   5080: 'Carrier 79 Drive: Short-circuit/ground fault detected', class No Acknowledgement, trigger "DB302_HMI_Faults_Carrier79_Faults_1" bit 7
   5081: 'Carrier 79 Drive: PROFINET Setpoint timeout', class No Acknowledgement, trigger "DB302_HMI_Faults_Carrier79_Faults_1" bit 8
   5082: 'Carrier 79 Power unit: Overcurrent', class No Acknowledgement, trigger "DB302_HMI_Faults_Carrier79_Faults_1" bit 9
   5083: 'Carrier 79 Power unit: DC link voltage overvoltage', class No Acknowledgement, trigger "DB302_HMI_Faults_Carrier79_Faults_1" bit 10
   5084: 'Carrier 79 Power unit: DC link voltage undervoltage', class No Acknowledgement, trigger "DB302_HMI_Faults_Carrier79_Faults_1" bit 11
   5085: 'Carrier 79 Power unit: Line phase failure in main circuit', class No Acknowledgement, trigger "DB302_HMI_Faults_Carrier79_Faults_1" bit 12
   5086: 'Carrier 79 Power unit: Phase failure motor cable', class No Acknowledgement, trigger "DB302_HMI_Faults_Carrier79_Faults_1" bit 13
   5087: 'Carrier 79 Power unit: Ground fault', class No Acknowledgement, trigger "DB302_HMI_Faults_Carrier79_Faults_1" bit 14
   5088: 'Spare_Fault_5088', class No Acknowledgement, trigger "DB302_HMI_Faults_Carrier79_Faults_1" bit 15
   5089: 'Carrier 79 Motion Off Fault', class No Acknowledgement, trigger "DB302_HMI_Faults_Carrier79_Faults_2" bit 0
   5090: 'Carrier 79 Motion On Fault', class No Acknowledgement, trigger "DB302_HMI_Faults_Carrier79_Faults_2" bit 1
   5091: 'Carrier 79 Spacing Fault', class No Acknowledgement, trigger "DB302_HMI_Faults_Carrier79_Faults_2" bit 2
   5092: 'Carrier 79 Duplicate Carrier Number Fault', class No Acknowledgement, trigger "DB302_HMI_Faults_Carrier79_Faults_2" bit 3
   5093: 'Spare_Fault_5093', class No Acknowledgement, trigger "DB302_HMI_Faults_Carrier79_Faults_2" bit 4
   5094: 'Spare_Fault_5094', class No Acknowledgement, trigger "DB302_HMI_Faults_Carrier79_Faults_2" bit 5
   5095: 'Spare_Fault_5095', class No Acknowledgement, trigger "DB302_HMI_Faults_Carrier79_Faults_2" bit 6
   5096: 'Spare_Fault_5096', class No Acknowledgement, trigger "DB302_HMI_Faults_Carrier79_Faults_2" bit 7
   5097: 'Spare_Fault_5097', class No Acknowledgement, trigger "DB302_HMI_Faults_Carrier79_Faults_2" bit 8
   5098: 'Spare_Fault_5098', class No Acknowledgement, trigger "DB302_HMI_Faults_Carrier79_Faults_2" bit 9
   5099: 'Spare_Fault_5099', class No Acknowledgement, trigger "DB302_HMI_Faults_Carrier79_Faults_2" bit 10
   5100: 'Spare_Fault_5100', class No Acknowledgement, trigger "DB302_HMI_Faults_Carrier79_Faults_2" bit 11
   5101: 'Spare_Fault_5101', class No Acknowledgement, trigger "DB302_HMI_Faults_Carrier79_Faults_2" bit 12
   5102: 'Spare_Fault_5102', class No Acknowledgement, trigger "DB302_HMI_Faults_Carrier79_Faults_2" bit 13
   5103: 'Spare_Fault_5103', class No Acknowledgement, trigger "DB302_HMI_Faults_Carrier79_Faults_2" bit 14
   5104: 'Spare_Fault_5104', class No Acknowledgement, trigger "DB302_HMI_Faults_Carrier79_Faults_2" bit 15
   5105: 'Spare_Fault_5105', class No Acknowledgement, trigger "DB302_HMI_Faults_Carrier79_Faults_3" bit 0
   5106: 'Spare_Fault_5106', class No Acknowledgement, trigger "DB302_HMI_Faults_Carrier79_Faults_3" bit 1
   5107: 'Spare_Fault_5107', class No Acknowledgement, trigger "DB302_HMI_Faults_Carrier79_Faults_3" bit 2
   5108: 'Spare_Fault_5108', class No Acknowledgement, trigger "DB302_HMI_Faults_Carrier79_Faults_3" bit 3
   5109: 'Spare_Fault_5109', class No Acknowledgement, trigger "DB302_HMI_Faults_Carrier79_Faults_3" bit 4
   5110: 'Spare_Fault_5110', class No Acknowledgement, trigger "DB302_HMI_Faults_Carrier79_Faults_3" bit 5
   5111: 'Spare_Fault_5111', class No Acknowledgement, trigger "DB302_HMI_Faults_Carrier79_Faults_3" bit 6
   5112: 'Spare_Fault_5112', class No Acknowledgement, trigger "DB302_HMI_Faults_Carrier79_Faults_3" bit 7
   5113: 'Spare_Fault_5113', class No Acknowledgement, trigger "DB302_HMI_Faults_Carrier79_Faults_3" bit 8
   5114: 'Spare_Fault_5114', class No Acknowledgement, trigger "DB302_HMI_Faults_Carrier79_Faults_3" bit 9
   5115: 'Spare_Fault_5115', class No Acknowledgement, trigger "DB302_HMI_Faults_Carrier79_Faults_3" bit 10
   5116: 'Spare_Fault_5116', class No Acknowledgement, trigger "DB302_HMI_Faults_Carrier79_Faults_3" bit 11
   5117: 'Spare_Fault_5117', class No Acknowledgement, trigger "DB302_HMI_Faults_Carrier79_Faults_3" bit 12
   5118: 'Spare_Fault_5118', class No Acknowledgement, trigger "DB302_HMI_Faults_Carrier79_Faults_3" bit 13
   5119: 'Spare_Fault_5119', class No Acknowledgement, trigger "DB302_HMI_Faults_Carrier79_Faults_3" bit 14
   5120: 'Spare_Fault_5120', class No Acknowledgement, trigger "DB302_HMI_Faults_Carrier79_Faults_3" bit 15
   5121: 'Carrier 80 Disconnect Open Power Fault DI11.0', class No Acknowledgement, trigger "DB302_HMI_Faults_Carrier80_Faults_0" bit 0
   5122: 'Carrier 80 Drive Profinet Comm Fault', class No Acknowledgement, trigger "DB302_HMI_Faults_Carrier80_Faults_0" bit 1
   5123: 'Carrier 80 Production Stop Not Reset', class No Acknowledgement, trigger "DB302_HMI_Faults_Carrier80_Faults_0" bit 2
   5124: 'Carrier 80 CB02122 Tripped', class No Acknowledgement, trigger "DB302_HMI_Faults_Carrier80_Faults_0" bit 3
   5125: 'Carrier 80 CB02123 Tripped', class No Acknowledgement, trigger "DB302_HMI_Faults_Carrier80_Faults_0" bit 4
   5126: 'Carrier 80 AUX1 CB Tripped', class No Acknowledgement, trigger "DB302_HMI_Faults_Carrier80_Faults_0" bit 5
   5127: 'Carrier 80 AUX2 CB Tripped', class No Acknowledgement, trigger "DB302_HMI_Faults_Carrier80_Faults_0" bit 6
   5128: 'Carrier 80 PLC Not Communicating', class No Acknowledgement, trigger "DB302_HMI_Faults_Carrier80_Faults_0" bit 7
   5129: 'Carrier 80 Safe Input Card Fault', class No Acknowledgement, trigger "DB302_HMI_Faults_Carrier80_Faults_0" bit 8
   5130: 'Carrier 80 Safe Output Card Fault', class No Acknowledgement, trigger "DB302_HMI_Faults_Carrier80_Faults_0" bit 9
   5131: 'Carrier 80 Standard Input Card Fault', class No Acknowledgement, trigger "DB302_HMI_Faults_Carrier80_Faults_0" bit 10
   5132: 'Carrier 80 Standard Output Card Fault', class No Acknowledgement, trigger "DB302_HMI_Faults_Carrier80_Faults_0" bit 11
   5133: 'Carrier 80 Encoder Position Fault', class No Acknowledgement, trigger "DB302_HMI_Faults_Carrier80_Faults_0" bit 12
   5134: 'Carrier 80 Encoder Internal Error', class No Acknowledgement, trigger "DB302_HMI_Faults_Carrier80_Faults_0" bit 13
   5135: 'Carrier 80 Encoder Comm Fault', class No Acknowledgement, trigger "DB302_HMI_Faults_Carrier80_Faults_0" bit 14
   5136: 'Carrier 80 HMI Comm Fault', class No Acknowledgement, trigger "DB302_HMI_Faults_Carrier80_Faults_0" bit 15
   5137: 'Carrier 80 Crash Detection Fault', class No Acknowledgement, trigger "DB302_HMI_Faults_Carrier80_Faults_1" bit 0
   5138: 'Carrier 80 Carrier Number Invalid', class No Acknowledgement, trigger "DB302_HMI_Faults_Carrier80_Faults_1" bit 1
   5139: 'Carrier 80 Drive: PROFINET configuration error', class No Acknowledgement, trigger "DB302_HMI_Faults_Carrier80_Faults_1" bit 2
   5140: 'Carrier 80 Drive: Error internal communications', class No Acknowledgement, trigger "DB302_HMI_Faults_Carrier80_Faults_1" bit 3
   5141: 'Carrier 80 Drive: Motor overtemperature', class No Acknowledgement, trigger "DB302_HMI_Faults_Carrier80_Faults_1" bit 4
   5142: 'Carrier 80 Drive: Motor overcurrent', class No Acknowledgement, trigger "DB302_HMI_Faults_Carrier80_Faults_1" bit 5
   5143: 'Carrier 80 Drive: Infeed or power unit not ready', class No Acknowledgement, trigger "DB302_HMI_Faults_Carrier80_Faults_1" bit 6
   5144: 'Carrier 80 Drive: Short-circuit/ground fault detected', class No Acknowledgement, trigger "DB302_HMI_Faults_Carrier80_Faults_1" bit 7
   5145: 'Carrier 80 Drive: PROFINET Setpoint timeout', class No Acknowledgement, trigger "DB302_HMI_Faults_Carrier80_Faults_1" bit 8
   5146: 'Carrier 80 Power unit: Overcurrent', class No Acknowledgement, trigger "DB302_HMI_Faults_Carrier80_Faults_1" bit 9
   5147: 'Carrier 80 Power unit: DC link voltage overvoltage', class No Acknowledgement, trigger "DB302_HMI_Faults_Carrier80_Faults_1" bit 10
   5148: 'Carrier 80 Power unit: DC link voltage undervoltage', class No Acknowledgement, trigger "DB302_HMI_Faults_Carrier80_Faults_1" bit 11
   5149: 'Carrier 80 Power unit: Line phase failure in main circuit', class No Acknowledgement, trigger "DB302_HMI_Faults_Carrier80_Faults_1" bit 12
   5150: 'Carrier 80 Power unit: Phase failure motor cable', class No Acknowledgement, trigger "DB302_HMI_Faults_Carrier80_Faults_1" bit 13
   5151: 'Carrier 80 Power unit: Ground fault', class No Acknowledgement, trigger "DB302_HMI_Faults_Carrier80_Faults_1" bit 14
   5152: 'Spare_Fault_5152', class No Acknowledgement, trigger "DB302_HMI_Faults_Carrier80_Faults_1" bit 15
   5153: 'Carrier 80 Motion Off Fault', class No Acknowledgement, trigger "DB302_HMI_Faults_Carrier80_Faults_2" bit 0
   5154: 'Carrier 80 Motion On Fault', class No Acknowledgement, trigger "DB302_HMI_Faults_Carrier80_Faults_2" bit 1
   5155: 'Carrier 80 Spacing Fault', class No Acknowledgement, trigger "DB302_HMI_Faults_Carrier80_Faults_2" bit 2
   5156: 'Carrier 80 Duplicate Carrier Number Fault', class No Acknowledgement, trigger "DB302_HMI_Faults_Carrier80_Faults_2" bit 3
   5157: 'Spare_Fault_5157', class No Acknowledgement, trigger "DB302_HMI_Faults_Carrier80_Faults_2" bit 4
   5158: 'Spare_Fault_5158', class No Acknowledgement, trigger "DB302_HMI_Faults_Carrier80_Faults_2" bit 5
   5159: 'Spare_Fault_5159', class No Acknowledgement, trigger "DB302_HMI_Faults_Carrier80_Faults_2" bit 6
   5160: 'Spare_Fault_5160', class No Acknowledgement, trigger "DB302_HMI_Faults_Carrier80_Faults_2" bit 7
   5161: 'Spare_Fault_5161', class No Acknowledgement, trigger "DB302_HMI_Faults_Carrier80_Faults_2" bit 8
   5162: 'Spare_Fault_5162', class No Acknowledgement, trigger "DB302_HMI_Faults_Carrier80_Faults_2" bit 9
   5163: 'Spare_Fault_5163', class No Acknowledgement, trigger "DB302_HMI_Faults_Carrier80_Faults_2" bit 10
   5164: 'Spare_Fault_5164', class No Acknowledgement, trigger "DB302_HMI_Faults_Carrier80_Faults_2" bit 11
   5165: 'Spare_Fault_5165', class No Acknowledgement, trigger "DB302_HMI_Faults_Carrier80_Faults_2" bit 12
   5166: 'Spare_Fault_5166', class No Acknowledgement, trigger "DB302_HMI_Faults_Carrier80_Faults_2" bit 13
   5167: 'Spare_Fault_5167', class No Acknowledgement, trigger "DB302_HMI_Faults_Carrier80_Faults_2" bit 14
   5168: 'Spare_Fault_5168', class No Acknowledgement, trigger "DB302_HMI_Faults_Carrier80_Faults_2" bit 15
   5169: 'Spare_Fault_5169', class No Acknowledgement, trigger "DB302_HMI_Faults_Carrier80_Faults_3" bit 0
   5170: 'Spare_Fault_5170', class No Acknowledgement, trigger "DB302_HMI_Faults_Carrier80_Faults_3" bit 1
   5171: 'Spare_Fault_5171', class No Acknowledgement, trigger "DB302_HMI_Faults_Carrier80_Faults_3" bit 2
   5172: 'Spare_Fault_5172', class No Acknowledgement, trigger "DB302_HMI_Faults_Carrier80_Faults_3" bit 3
   5173: 'Spare_Fault_5173', class No Acknowledgement, trigger "DB302_HMI_Faults_Carrier80_Faults_3" bit 4
   5174: 'Spare_Fault_5174', class No Acknowledgement, trigger "DB302_HMI_Faults_Carrier80_Faults_3" bit 5
   5175: 'Spare_Fault_5175', class No Acknowledgement, trigger "DB302_HMI_Faults_Carrier80_Faults_3" bit 6
   5176: 'Spare_Fault_5176', class No Acknowledgement, trigger "DB302_HMI_Faults_Carrier80_Faults_3" bit 7
   5177: 'Spare_Fault_5177', class No Acknowledgement, trigger "DB302_HMI_Faults_Carrier80_Faults_3" bit 8
   5178: 'Spare_Fault_5178', class No Acknowledgement, trigger "DB302_HMI_Faults_Carrier80_Faults_3" bit 9
   5179: 'Spare_Fault_5179', class No Acknowledgement, trigger "DB302_HMI_Faults_Carrier80_Faults_3" bit 10
   5180: 'Spare_Fault_5180', class No Acknowledgement, trigger "DB302_HMI_Faults_Carrier80_Faults_3" bit 11
   5181: 'Spare_Fault_5181', class No Acknowledgement, trigger "DB302_HMI_Faults_Carrier80_Faults_3" bit 12
   5182: 'Spare_Fault_5182', class No Acknowledgement, trigger "DB302_HMI_Faults_Carrier80_Faults_3" bit 13
   5183: 'Spare_Fault_5183', class No Acknowledgement, trigger "DB302_HMI_Faults_Carrier80_Faults_3" bit 14
   5184: 'Spare_Fault_5184', class No Acknowledgement, trigger "DB302_HMI_Faults_Carrier80_Faults_3" bit 15
   5185: 'Carrier 81 Disconnect Open Power Fault DI11.0', class No Acknowledgement, trigger "DB302_HMI_Faults_Carrier81_Faults_0" bit 0
   5186: 'Carrier 81 Drive Profinet Comm Fault', class No Acknowledgement, trigger "DB302_HMI_Faults_Carrier81_Faults_0" bit 1
   5187: 'Carrier 81 Production Stop Not Reset', class No Acknowledgement, trigger "DB302_HMI_Faults_Carrier81_Faults_0" bit 2
   5188: 'Carrier 81 CB02122 Tripped', class No Acknowledgement, trigger "DB302_HMI_Faults_Carrier81_Faults_0" bit 3
   5189: 'Carrier 81 CB02123 Tripped', class No Acknowledgement, trigger "DB302_HMI_Faults_Carrier81_Faults_0" bit 4
   5190: 'Carrier 81 AUX1 CB Tripped', class No Acknowledgement, trigger "DB302_HMI_Faults_Carrier81_Faults_0" bit 5
   5191: 'Carrier 81 AUX2 CB Tripped', class No Acknowledgement, trigger "DB302_HMI_Faults_Carrier81_Faults_0" bit 6
   5192: 'Carrier 81 PLC Not Communicating', class No Acknowledgement, trigger "DB302_HMI_Faults_Carrier81_Faults_0" bit 7
   5193: 'Carrier 81 Safe Input Card Fault', class No Acknowledgement, trigger "DB302_HMI_Faults_Carrier81_Faults_0" bit 8
   5194: 'Carrier 81 Safe Output Card Fault', class No Acknowledgement, trigger "DB302_HMI_Faults_Carrier81_Faults_0" bit 9
   5195: 'Carrier 81 Standard Input Card Fault', class No Acknowledgement, trigger "DB302_HMI_Faults_Carrier81_Faults_0" bit 10
   5196: 'Carrier 81 Standard Output Card Fault', class No Acknowledgement, trigger "DB302_HMI_Faults_Carrier81_Faults_0" bit 11
   5197: 'Carrier 81 Encoder Position Fault', class No Acknowledgement, trigger "DB302_HMI_Faults_Carrier81_Faults_0" bit 12
   5198: 'Carrier 81 Encoder Internal Error', class No Acknowledgement, trigger "DB302_HMI_Faults_Carrier81_Faults_0" bit 13
   5199: 'Carrier 81 Encoder Comm Fault', class No Acknowledgement, trigger "DB302_HMI_Faults_Carrier81_Faults_0" bit 14
   5200: 'Carrier 81 HMI Comm Fault', class No Acknowledgement, trigger "DB302_HMI_Faults_Carrier81_Faults_0" bit 15
   5201: 'Carrier 81 Crash Detection Fault', class No Acknowledgement, trigger "DB302_HMI_Faults_Carrier81_Faults_1" bit 0
   5202: 'Carrier 81 Carrier Number Invalid', class No Acknowledgement, trigger "DB302_HMI_Faults_Carrier81_Faults_1" bit 1
   5203: 'Carrier 81 Drive: PROFINET configuration error', class No Acknowledgement, trigger "DB302_HMI_Faults_Carrier81_Faults_1" bit 2
   5204: 'Carrier 81 Drive: Error internal communications', class No Acknowledgement, trigger "DB302_HMI_Faults_Carrier81_Faults_1" bit 3
   5205: 'Carrier 81 Drive: Motor overtemperature', class No Acknowledgement, trigger "DB302_HMI_Faults_Carrier81_Faults_1" bit 4
   5206: 'Carrier 81 Drive: Motor overcurrent', class No Acknowledgement, trigger "DB302_HMI_Faults_Carrier81_Faults_1" bit 5
   5207: 'Carrier 81 Drive: Infeed or power unit not ready', class No Acknowledgement, trigger "DB302_HMI_Faults_Carrier81_Faults_1" bit 6
   5208: 'Carrier 81 Drive: Short-circuit/ground fault detected', class No Acknowledgement, trigger "DB302_HMI_Faults_Carrier81_Faults_1" bit 7
   5209: 'Carrier 81 Drive: PROFINET Setpoint timeout', class No Acknowledgement, trigger "DB302_HMI_Faults_Carrier81_Faults_1" bit 8
   5210: 'Carrier 81 Power unit: Overcurrent', class No Acknowledgement, trigger "DB302_HMI_Faults_Carrier81_Faults_1" bit 9
   5211: 'Carrier 81 Power unit: DC link voltage overvoltage', class No Acknowledgement, trigger "DB302_HMI_Faults_Carrier81_Faults_1" bit 10
   5212: 'Carrier 81 Power unit: DC link voltage undervoltage', class No Acknowledgement, trigger "DB302_HMI_Faults_Carrier81_Faults_1" bit 11
   5213: 'Carrier 81 Power unit: Line phase failure in main circuit', class No Acknowledgement, trigger "DB302_HMI_Faults_Carrier81_Faults_1" bit 12
   5214: 'Carrier 81 Power unit: Phase failure motor cable', class No Acknowledgement, trigger "DB302_HMI_Faults_Carrier81_Faults_1" bit 13
   5215: 'Carrier 81 Power unit: Ground fault', class No Acknowledgement, trigger "DB302_HMI_Faults_Carrier81_Faults_1" bit 14
   5216: 'Spare_Fault_5216', class No Acknowledgement, trigger "DB302_HMI_Faults_Carrier81_Faults_1" bit 15
   5217: 'Carrier 81 Motion Off Fault', class No Acknowledgement, trigger "DB302_HMI_Faults_Carrier81_Faults_2" bit 0
   5218: 'Carrier 81 Motion On Fault', class No Acknowledgement, trigger "DB302_HMI_Faults_Carrier81_Faults_2" bit 1
   5219: 'Carrier 81 Spacing Fault', class No Acknowledgement, trigger "DB302_HMI_Faults_Carrier81_Faults_2" bit 2
   5220: 'Carrier 81 Duplicate Carrier Number Fault', class No Acknowledgement, trigger "DB302_HMI_Faults_Carrier81_Faults_2" bit 3
   5221: 'Spare_Fault_5221', class No Acknowledgement, trigger "DB302_HMI_Faults_Carrier81_Faults_2" bit 4
   5222: 'Spare_Fault_5222', class No Acknowledgement, trigger "DB302_HMI_Faults_Carrier81_Faults_2" bit 5
   5223: 'Spare_Fault_5223', class No Acknowledgement, trigger "DB302_HMI_Faults_Carrier81_Faults_2" bit 6
   5224: 'Spare_Fault_5224', class No Acknowledgement, trigger "DB302_HMI_Faults_Carrier81_Faults_2" bit 7
   5225: 'Spare_Fault_5225', class No Acknowledgement, trigger "DB302_HMI_Faults_Carrier81_Faults_2" bit 8
   5226: 'Spare_Fault_5226', class No Acknowledgement, trigger "DB302_HMI_Faults_Carrier81_Faults_2" bit 9
   5227: 'Spare_Fault_5227', class No Acknowledgement, trigger "DB302_HMI_Faults_Carrier81_Faults_2" bit 10
   5228: 'Spare_Fault_5228', class No Acknowledgement, trigger "DB302_HMI_Faults_Carrier81_Faults_2" bit 11
   5229: 'Spare_Fault_5229', class No Acknowledgement, trigger "DB302_HMI_Faults_Carrier81_Faults_2" bit 12
   5230: 'Spare_Fault_5230', class No Acknowledgement, trigger "DB302_HMI_Faults_Carrier81_Faults_2" bit 13
   5231: 'Spare_Fault_5231', class No Acknowledgement, trigger "DB302_HMI_Faults_Carrier81_Faults_2" bit 14
   5232: 'Spare_Fault_5232', class No Acknowledgement, trigger "DB302_HMI_Faults_Carrier81_Faults_2" bit 15
   5233: 'Spare_Fault_5233', class No Acknowledgement, trigger "DB302_HMI_Faults_Carrier81_Faults_3" bit 0
   5234: 'Spare_Fault_5234', class No Acknowledgement, trigger "DB302_HMI_Faults_Carrier81_Faults_3" bit 1
   5235: 'Spare_Fault_5235', class No Acknowledgement, trigger "DB302_HMI_Faults_Carrier81_Faults_3" bit 2
   5236: 'Spare_Fault_5236', class No Acknowledgement, trigger "DB302_HMI_Faults_Carrier81_Faults_3" bit 3
   5237: 'Spare_Fault_5237', class No Acknowledgement, trigger "DB302_HMI_Faults_Carrier81_Faults_3" bit 4
   5238: 'Spare_Fault_5238', class No Acknowledgement, trigger "DB302_HMI_Faults_Carrier81_Faults_3" bit 5
   5239: 'Spare_Fault_5239', class No Acknowledgement, trigger "DB302_HMI_Faults_Carrier81_Faults_3" bit 6
   5240: 'Spare_Fault_5240', class No Acknowledgement, trigger "DB302_HMI_Faults_Carrier81_Faults_3" bit 7
   5241: 'Spare_Fault_5241', class No Acknowledgement, trigger "DB302_HMI_Faults_Carrier81_Faults_3" bit 8
   5242: 'Spare_Fault_5242', class No Acknowledgement, trigger "DB302_HMI_Faults_Carrier81_Faults_3" bit 9
   5243: 'Spare_Fault_5243', class No Acknowledgement, trigger "DB302_HMI_Faults_Carrier81_Faults_3" bit 10
   5244: 'Spare_Fault_5244', class No Acknowledgement, trigger "DB302_HMI_Faults_Carrier81_Faults_3" bit 11
   5245: 'Spare_Fault_5245', class No Acknowledgement, trigger "DB302_HMI_Faults_Carrier81_Faults_3" bit 12
   5246: 'Spare_Fault_5246', class No Acknowledgement, trigger "DB302_HMI_Faults_Carrier81_Faults_3" bit 13
   5247: 'Spare_Fault_5247', class No Acknowledgement, trigger "DB302_HMI_Faults_Carrier81_Faults_3" bit 14
   5248: 'Spare_Fault_5248', class No Acknowledgement, trigger "DB302_HMI_Faults_Carrier81_Faults_3" bit 15
   5249: 'Carrier 82 Disconnect Open Power Fault DI11.0', class No Acknowledgement, trigger "DB302_HMI_Faults_Carrier82_Faults_0" bit 0
   5250: 'Carrier 82 Drive Profinet Comm Fault', class No Acknowledgement, trigger "DB302_HMI_Faults_Carrier82_Faults_0" bit 1
   5251: 'Carrier 82 Production Stop Not Reset', class No Acknowledgement, trigger "DB302_HMI_Faults_Carrier82_Faults_0" bit 2
   5252: 'Carrier 82 CB02122 Tripped', class No Acknowledgement, trigger "DB302_HMI_Faults_Carrier82_Faults_0" bit 3
   5253: 'Carrier 82 CB02123 Tripped', class No Acknowledgement, trigger "DB302_HMI_Faults_Carrier82_Faults_0" bit 4
   5254: 'Carrier 82 AUX1 CB Tripped', class No Acknowledgement, trigger "DB302_HMI_Faults_Carrier82_Faults_0" bit 5
   5255: 'Carrier 82 AUX2 CB Tripped', class No Acknowledgement, trigger "DB302_HMI_Faults_Carrier82_Faults_0" bit 6
   5256: 'Carrier 82 PLC Not Communicating', class No Acknowledgement, trigger "DB302_HMI_Faults_Carrier82_Faults_0" bit 7
   5257: 'Carrier 82 Safe Input Card Fault', class No Acknowledgement, trigger "DB302_HMI_Faults_Carrier82_Faults_0" bit 8
   5258: 'Carrier 82 Safe Output Card Fault', class No Acknowledgement, trigger "DB302_HMI_Faults_Carrier82_Faults_0" bit 9
   5259: 'Carrier 82 Standard Input Card Fault', class No Acknowledgement, trigger "DB302_HMI_Faults_Carrier82_Faults_0" bit 10
   5260: 'Carrier 82 Standard Output Card Fault', class No Acknowledgement, trigger "DB302_HMI_Faults_Carrier82_Faults_0" bit 11
   5261: 'Carrier 82 Encoder Position Fault', class No Acknowledgement, trigger "DB302_HMI_Faults_Carrier82_Faults_0" bit 12
   5262: 'Carrier 82 Encoder Internal Error', class No Acknowledgement, trigger "DB302_HMI_Faults_Carrier82_Faults_0" bit 13
   5263: 'Carrier 82 Encoder Comm Fault', class No Acknowledgement, trigger "DB302_HMI_Faults_Carrier82_Faults_0" bit 14
   5264: 'Carrier 82 HMI Comm Fault', class No Acknowledgement, trigger "DB302_HMI_Faults_Carrier82_Faults_0" bit 15
   5265: 'Carrier 82 Crash Detection Fault', class No Acknowledgement, trigger "DB302_HMI_Faults_Carrier82_Faults_1" bit 0
   5266: 'Carrier 82 Carrier Number Invalid', class No Acknowledgement, trigger "DB302_HMI_Faults_Carrier82_Faults_1" bit 1
   5267: 'Carrier 82 Drive: PROFINET configuration error', class No Acknowledgement, trigger "DB302_HMI_Faults_Carrier82_Faults_1" bit 2
   5268: 'Carrier 82 Drive: Error internal communications', class No Acknowledgement, trigger "DB302_HMI_Faults_Carrier82_Faults_1" bit 3
   5269: 'Carrier 82 Drive: Motor overtemperature', class No Acknowledgement, trigger "DB302_HMI_Faults_Carrier82_Faults_1" bit 4
   5270: 'Carrier 82 Drive: Motor overcurrent', class No Acknowledgement, trigger "DB302_HMI_Faults_Carrier82_Faults_1" bit 5
   5271: 'Carrier 82 Drive: Infeed or power unit not ready', class No Acknowledgement, trigger "DB302_HMI_Faults_Carrier82_Faults_1" bit 6
   5272: 'Carrier 82 Drive: Short-circuit/ground fault detected', class No Acknowledgement, trigger "DB302_HMI_Faults_Carrier82_Faults_1" bit 7
   5273: 'Carrier 82 Drive: PROFINET Setpoint timeout', class No Acknowledgement, trigger "DB302_HMI_Faults_Carrier82_Faults_1" bit 8
   5274: 'Carrier 82 Power unit: Overcurrent', class No Acknowledgement, trigger "DB302_HMI_Faults_Carrier82_Faults_1" bit 9
   5275: 'Carrier 82 Power unit: DC link voltage overvoltage', class No Acknowledgement, trigger "DB302_HMI_Faults_Carrier82_Faults_1" bit 10
   5276: 'Carrier 82 Power unit: DC link voltage undervoltage', class No Acknowledgement, trigger "DB302_HMI_Faults_Carrier82_Faults_1" bit 11
   5277: 'Carrier 82 Power unit: Line phase failure in main circuit', class No Acknowledgement, trigger "DB302_HMI_Faults_Carrier82_Faults_1" bit 12
   5278: 'Carrier 82 Power unit: Phase failure motor cable', class No Acknowledgement, trigger "DB302_HMI_Faults_Carrier82_Faults_1" bit 13
   5279: 'Carrier 82 Power unit: Ground fault', class No Acknowledgement, trigger "DB302_HMI_Faults_Carrier82_Faults_1" bit 14
   5280: 'Spare_Fault_5280', class No Acknowledgement, trigger "DB302_HMI_Faults_Carrier82_Faults_1" bit 15
   5281: 'Carrier 82 Motion Off Fault', class No Acknowledgement, trigger "DB302_HMI_Faults_Carrier82_Faults_2" bit 0
   5282: 'Carrier 82 Motion On Fault', class No Acknowledgement, trigger "DB302_HMI_Faults_Carrier82_Faults_2" bit 1
   5283: 'Carrier 82 Spacing Fault', class No Acknowledgement, trigger "DB302_HMI_Faults_Carrier82_Faults_2" bit 2
   5284: 'Carrier 82 Duplicate Carrier Number Fault', class No Acknowledgement, trigger "DB302_HMI_Faults_Carrier82_Faults_2" bit 3
   5285: 'Spare_Fault_5285', class No Acknowledgement, trigger "DB302_HMI_Faults_Carrier82_Faults_2" bit 4
   5286: 'Spare_Fault_5286', class No Acknowledgement, trigger "DB302_HMI_Faults_Carrier82_Faults_2" bit 5
   5287: 'Spare_Fault_5287', class No Acknowledgement, trigger "DB302_HMI_Faults_Carrier82_Faults_2" bit 6
   5288: 'Spare_Fault_5288', class No Acknowledgement, trigger "DB302_HMI_Faults_Carrier82_Faults_2" bit 7
   5289: 'Spare_Fault_5289', class No Acknowledgement, trigger "DB302_HMI_Faults_Carrier82_Faults_2" bit 8
   5290: 'Spare_Fault_5290', class No Acknowledgement, trigger "DB302_HMI_Faults_Carrier82_Faults_2" bit 9
   5291: 'Spare_Fault_5291', class No Acknowledgement, trigger "DB302_HMI_Faults_Carrier82_Faults_2" bit 10
   5292: 'Spare_Fault_5292', class No Acknowledgement, trigger "DB302_HMI_Faults_Carrier82_Faults_2" bit 11
   5293: 'Spare_Fault_5293', class No Acknowledgement, trigger "DB302_HMI_Faults_Carrier82_Faults_2" bit 12
   5294: 'Spare_Fault_5294', class No Acknowledgement, trigger "DB302_HMI_Faults_Carrier82_Faults_2" bit 13
   5295: 'Spare_Fault_5295', class No Acknowledgement, trigger "DB302_HMI_Faults_Carrier82_Faults_2" bit 14
   5296: 'Spare_Fault_5296', class No Acknowledgement, trigger "DB302_HMI_Faults_Carrier82_Faults_2" bit 15
   5297: 'Spare_Fault_5297', class No Acknowledgement, trigger "DB302_HMI_Faults_Carrier82_Faults_3" bit 0
   5298: 'Spare_Fault_5298', class No Acknowledgement, trigger "DB302_HMI_Faults_Carrier82_Faults_3" bit 1
   5299: 'Spare_Fault_5299', class No Acknowledgement, trigger "DB302_HMI_Faults_Carrier82_Faults_3" bit 2
   5300: 'Spare_Fault_5300', class No Acknowledgement, trigger "DB302_HMI_Faults_Carrier82_Faults_3" bit 3
   5301: 'Spare_Fault_5301', class No Acknowledgement, trigger "DB302_HMI_Faults_Carrier82_Faults_3" bit 4
   5302: 'Spare_Fault_5302', class No Acknowledgement, trigger "DB302_HMI_Faults_Carrier82_Faults_3" bit 5
   5303: 'Spare_Fault_5303', class No Acknowledgement, trigger "DB302_HMI_Faults_Carrier82_Faults_3" bit 6
   5304: 'Spare_Fault_5304', class No Acknowledgement, trigger "DB302_HMI_Faults_Carrier82_Faults_3" bit 7
   5305: 'Spare_Fault_5305', class No Acknowledgement, trigger "DB302_HMI_Faults_Carrier82_Faults_3" bit 8
   5306: 'Spare_Fault_5306', class No Acknowledgement, trigger "DB302_HMI_Faults_Carrier82_Faults_3" bit 9
   5307: 'Spare_Fault_5307', class No Acknowledgement, trigger "DB302_HMI_Faults_Carrier82_Faults_3" bit 10
   5308: 'Spare_Fault_5308', class No Acknowledgement, trigger "DB302_HMI_Faults_Carrier82_Faults_3" bit 11
   5309: 'Spare_Fault_5309', class No Acknowledgement, trigger "DB302_HMI_Faults_Carrier82_Faults_3" bit 12
   5310: 'Spare_Fault_5310', class No Acknowledgement, trigger "DB302_HMI_Faults_Carrier82_Faults_3" bit 13
   5311: 'Spare_Fault_5311', class No Acknowledgement, trigger "DB302_HMI_Faults_Carrier82_Faults_3" bit 14
   5312: 'Spare_Fault_5312', class No Acknowledgement, trigger "DB302_HMI_Faults_Carrier82_Faults_3" bit 15
   4: 'Wireless Access Point 3 Comm Fault', class No Acknowledgement, trigger "DB302_HMI_Faults_SDC_Faults_0" bit 3

text list "SDC_G120D": 0 ''; 0 'Antrieb hat keine Störung / kein Fehlercode'; 1000 'Softwarefehler intern'; 1001 'FloatingPoint Ausnahme'; 1002 'Softwarefehler intern'; 1003 'Quittungsverzug bei Speicherzugriff'; 1004 'Softwarefehler intern'; 1005 'Datei Upload/Download fehlgeschlagen'; 1009 'CU: Regelungsbaugruppe Übertemperatur'; 1010 'Antriebstyp unbekannt'; 1015 'Softwarefehler intern'; 1016 'Firmware verändert'; 1017 'Komponentenlisten verändert'; 1018 'Hochlauf mehrmals abgebrochen'; 1019 'Wechselmedium schreiben fehlgeschlagen'; 1020 'RAM disk Schreiben fehlgeschlagen'; 1021 'Wechselmedium als USB-Datenträger von PC verwendet'; 1023 'Software Timeout intern'; 1028 'Konfigurationsfehler'; 1030 'Lebenszeichenausfall bei Steuerungshoheit'; 1033 'Einheitenumschaltung: Bezugsparameterwert ungültig'; 1034 'Einheitenumschaltung: Berechnung Parameterwerte nach Bezugswertänderung fehlgeschlagen'; 1035 'ACX: Parametersicherungsdateien beschädigt'; 1036 'ACX: Parametersicherungsdatei fehlt'; 1038 'ACX: Parametersicherungsdatei laden fehlgeschlagen'; 1039 'ACX: Parametersicherungsdatei schreiben fehlgeschlagen'; 1040 'Parameter sichern und POWER ON erforderlich'; 1042 'Parameterfehler beim Projekt-Download'; 1043 'Schwerer Fehler beim Projekt-Download'; 1044 'CU: Beschreibungsdaten fehlerhaft'; 1045 'Projektierungsdaten ungültig'; 1049 'Schreiben in Datei nicht möglich'; 1054 'CU: Systemgrenze überschritten'; 1064 'CU: Interner Fehler (CRC)'; 1066 'Zwischenspeicher: Füllstand 70 % erreicht oder überschritten'; 1067 'Zwischenspeicher: Füllstand 100 % erreicht'; 1068 'CU: Datenspeicher Speicherüberlauf'; 1069 'Parametersicherung und Gerät inkompatibel'; 1072 'Speicherkarte aus Sicherungskopie wieder hergestellt'; 1073 'POWER ON für Sicherungskopie auf Speicherkarte erforderlich'; 1105 'CU: Speicher nicht ausreichend'; 1107 'Speichern auf Speicherkarte fehlgeschlagen'; 1112 'CU: Leistungsteil unzulässig'; 1120 'Initialisierung Klemmen fehlgeschlagen'; 1122 'Frequenz am Messtastereingang zu hoch'; 1205 'CU: Zeitscheibenüberlauf'; 1250 'CU: CU-EEPROM Read-Only-Daten fehlerhaft'; 1251 'CU: CU-EEPROM Read-Write-Daten fehlerhaft'; 1257 'CU: Firmware-Version veraltet'; 1340 'Topologie: Zu viele Komponenten an einem Strang'; 1505 'BICO: Verschaltung kann nicht hergestellt werden'; 1510 'BICO: Signalquelle ist nicht Float'; 1511 'BICO: Verschaltung mit unterschiedlicher Normierung'; 1512 'BICO: Keine Normierung vorhanden'; 1513 'BICO: Verschaltung DO-übergreifend mit unterschiedlicher Normierung'; 1514 'BICO: Fehler beim Schreiben während Reconnect'; 1515 'BICO: Parameterschreiben nicht erlaubt da Steuerungshoheit aktiv'; 1590 'Antrieb: Motor Wartungsintervall abgelaufen'; 1600 'SI P1: STOP A ausgelöst'; 1611 'SI P1: Defekt in einem Überwachungskanal'; 1620 'SI P1: Sicher abgeschaltetes Moment aktiv'; 1625 'SI P1: Lebenszeichen in Safety-Daten fehlerhaft'; 1649 'SI P1: Softwarefehler intern'; 1650 'SI P1: Abnahmetest erforderlich'; 1651 'SI P1: Synchronisation Safety-Zeitscheiben fehlgeschlagen'; 1653 'SI P1: PROFIBUS/PROFINET-Projektierung fehlerhaft'; 1654 'SI P1: PROFIsafe-Projektierung abweichend'; 1655 'SI P1: Abgleich der Überwachungsfunktionen'; 1656 'SI P1: Parameter Prozessor 2 fehlerhaft'; 1658 'SI P1: PROFIsafe-Telegrammnummer ungeeignet'; 1659 'SI P1: Schreibauftrag für Parameter abgewiesen'; 1660 'SI P1: Sichere Funktionen nicht unterstützt'; 1661 'SI P1: Simulation der Safety Eingänge aktiv'; 1662 'Fehler interne Kommunikation'; 1663 'SI P1: Kopieren der SI-Parameter abgelehnt'; 1665 'SI P1: System ist defekt'; 1666 'SI Motion P1: Statisches 1-Signal am F-DI für sichere Quittierung'; 1669 'SI Motion: Kombination von Motor und Leistungsteil ungünstig'; 1680 'SI Motion P1: Prüfsummenfehler sichere Überwachungen'; 1681 'SI Motion P1: Parameterwert falsch'; 1682 'SI Motion P1: Überwachungsfunktion nicht unterstützt'; 1683 'SI Motion P1: SLS-Freigabe fehlt'; 1690 'SI Motion: Datensicherungsproblem beim NVRAM'; 1692 'SI Motion P1: Parameterwert geberlos unzulässig'; 1693 'SI Motion P1: Safety-Parametrierung geändert POWER ON erforderlich'; 1696 'SI Motion: Testanwahl der Bewegungsüberwachungen im Hochlauf'; 1697 'SI Motion: Test der Bewegungsüberwachungen erforderlich'; 1698 'SI P1: Inbetriebnahmemodus aktiv'; 1699 'SI P1: Test der Abschaltpfade erforderlich'; 1700 'SI Motion P1: STOP A ausgelöst'; 1701 'SI Motion P1: STOP B ausgelöst'; 1706 'SI Motion P1: SAM/SBR Grenze überschritten'; 1711 'SI Motion P1: Defekt in einem Überwachungskanal'; 1712 'SI Motion P1: Defekt bei F-IO-Verarbeitung'; 1714 'SI Motion P1: Sicher begrenzte Geschwindigkeit überschritten'; 1716 'SI Motion P1: Toleranz für sichere Bewegungsrichtung überschritten'; 1770 'SI Motion P1: Diskrepanzfehler der fehlersicheren Eingänge'; 1772 'SI Motion P1: Teststop fehlersichere Eingänge/Ausgänge aktiv'; 1773 'SI Motion P1: Teststop fehlerhaft'; 1774 'SI Motion P1: Teststop notwendig'; 1796 'SI P1: Warten auf Kommunikation'; 1798 'SI Motion P1: Teststop läuft'; 1799 'SI Motion P1: Abnahmetestmodus aktiv'; 1900 'PROFIBUS: Konfigurationstelegramm fehlerhaft'; 1910 'Feldbus SS Sollwert Timeout'; 1920 'PROFIBUS: Unterbrechung zyklische Verbindung'; 1945 'PROFIBUS: Verbindung zum Publisher gestört'; 1946 'PROFIBUS: Verbindung zum Publisher abgebrochen'; 1951 'CU SYNC: Synchronisation Applikationstakt fehlt'; 1953 'CU SYNC: Synchronisation nicht abgeschlossen'; 2050 'Trace: Start nicht möglich'; 2055 'Trace: Aufzeichnungsdauer zu klein'; 2056 'Trace: Aufzeichnungstakt zu klein'; 2057 'Trace: Zeitscheibentakt ungültig'; 2058 'Trace: Zeitscheibentakt für Endlostrace ungültig'; 2059 'Trace: Zeitscheibentakt für 2 x 8 Aufzeichnungskanäle ungültig'; 2060 'Trace: Aufzuzeichnendes Signal fehlt'; 2061 'Trace: Signal ungültig'; 2062 'Trace: Triggersignal ungültig'; 2063 'Trace: Datentyp ungültig'; 2070 'Trace: Parameter nicht änderbar'; 2075 'Trace: Pretriggerzeit zu groß'; 2080 'Trace: Parametrierung wegen Einheitenumschaltung gelöscht'; 2097 'MTrace: Mehrfachtrace aktivieren nicht möglich'; 2098 'MTrace: Speichern nicht möglich'; 2099 'Trace: Speicherplatz der Control Unit nicht ausreichend'; 2150 'OA: Applikation nicht ladbar'; 2151 'OA: Softwarefehler intern'; 2152 'OA: Speicher nicht ausreichend'; 3000 'NVRAM Fehler bei Aktion'; 3001 'NVRAM Prüfsumme fehlerhaft'; 3505 'CU: Analogeingang Drahtbruch'; 3510 'CU: Kalibrierdaten nicht plausibel'; 5000 'Leistungsteil: Übertemperatur Kühlkörper Wechselrichter'; 5001 'Leistungsteil: Übertemperatur Sperrschicht Chip'; 5002 'Leistungsteil: Übertemperatur Zuluft'; 5004 'Leistungsteil: Übertemperatur Gleichrichter'; 5006 'Leistungsteil: Übertemperatur Thermisches Modell'; 6310 'Anschlussspannung (p0210) fehlerhaft parametriert'; 6921 'Bremswiderstand Phasenunsymmetrie'; 6922 'Bremswiderstand Phasenausfall'; 7011 'Antrieb: Motor Übertemperatur'; 7012 'Antrieb: Motortemperaturmodell 1 Übertemperatur'; 7014 'Antrieb: Motortemperaturmodell Konfiguration Warnung'; 7015 'Antrieb: Motortemperatursensor Warnung'; 7016 'Antrieb: Motortemperatursensor Störung'; 7080 'Antrieb: Regelungsparameter fehlerhaft'; 7082 'Makro: Ausführung nicht möglich'; 7083 'Makro: ACX-File nicht gefunden'; 7084 'Makro: Bedingung für WaitUntil nicht erfüllt'; 7086 'Einheitenumschaltung: Parametergrenzverletzung durch Bezugswertänderung'; 7088 'Einheitenumschaltung: Parametergrenzverletzung durch Einheitenumschaltung'; 7089 'Einheitenumschaltung: Funktionsmodul aktivieren ist blockiert weil Einheiten umgeschaltet'; 7200 'Antrieb: Steuerungshoheit EIN-Befehl steht an'; 7220 'Antrieb: Führung durch PLC fehlt'; 7300 'Antrieb: Netzschütz Rückmeldung fehlt'; 7320 'Antrieb: Automatischer Wiederanlauf abgebrochen'; 7321 'Antrieb: Automatischer Wiederanlauf aktiv'; 7330 'Fangen: Gemessener Suchstrom zu klein'; 7331 'Fangen: Funktion nicht unterstützt'; 7400 'Antrieb: Zwischenkreisspannungs-Maximum-Regler aktiv'; 7401 'Antrieb: Zwischenkreisspannungs-Maximum-Regler deaktiviert'; 7402 'Antrieb: Zwischenkreisspannungs-Minimum-Regler aktiv'; 7404 'Antrieb: Zwischenkreisspannungsüberwachnung Vdc_Max'; 7405 'Antrieb: Kinetische Pufferung minimale Drehzahl unterschritten'; 7406 'Antrieb: Kinetische Pufferung maximale Dauer überschritten'; 7409 'Antrieb: U/f-Steuerung Strombegrenzungsregler aktiv'; 7410 'Antrieb: Stromreglerausgang begrenzt'; 7411 'Antrieb: Flussreglerausgang begrenzt'; 7416 'Antrieb: Konfiguration Flussregler'; 7426 'Technologieregler Istwert begrenzt'; 7428 'Technologieregler Parametrierfehler'; 7435 'Antrieb: Hochlaufgebersetzen bei geberloser Vektorregelung'; 7440 'EPOS: Ruckzeit wird begrenzt'; 7441 'LR: Lageoffset der Absolutwertgeberjustage sichern'; 7442 'LR: Multiturn passt nicht zum Modulobereich'; 7443 'LR: Referenzpunkt-Koordinate nicht im zulässigen Bereich'; 7450 'LR: Stillstandsüberwachung hat angesprochen'; 7451 'LR: Positionierüberwachung hat angesprochen'; 7452 'LR: Schleppabstand zu groß'; 7453 'LR: Lageistwertaufbereitung fehlerhaft'; 7454 'LR: Lageistwertaufbereitung hat keinen gültigen Geber'; 7455 'EPOS: Maximalgeschwindigkeit begrenzt'; 7456 'EPOS: Sollgeschwindigkeit begrenzt'; 7457 'EPOS: Eingangssignale Kombination unzulässig'; 7458 'EPOS: Referenznocken nicht gefunden'; 7459 'EPOS: Keine Nullmarke vorhanden'; 7460 'EPOS: Referenznockenende nicht gefunden'; 7461 'EPOS: Referenzpunkt nicht gesetzt'; 7462 'EPOS: Angewählte Verfahrsatznummer existiert nicht'; 7463 'EPOS: Externer Satzwechsel im Verfahrsatz nicht angefordert'; 7464 'EPOS: Verfahrsatz ist inkonsistent'; 7465 'EPOS: Verfahrsatz hat keinen Folgesatz'; 7466 'EPOS: Verfahrsatznummer mehrfach vergeben'; 7467 'EPOS: Verfahrsatz hat unzulässigen Auftragsparameter'; 7468 'EPOS: Verfahrsatz Sprungziel existiert nicht'; 7469 'EPOS: Verfahrsatz Zielposition < Software-Endschalter Minus'; 7470 'EPOS: Verfahrsatz Zielposition > Software-Endschalter Plus'; 7471 'EPOS: Verfahrsatz Zielposition außerhalb Modulobereich'; 7472 'EPOS: Verfahrsatz ABS_POS/ABS_NEG nicht möglich'; 7473 'EPOS: Verfahrbereichsanfang angefahren'; 7474 'EPOS: Verfahrbereichsende angefahren'; 7475 'EPOS: Zielposition < Verfahrbereichsanfang'; 7476 'EPOS: Zielposition > Verfahrbereichsende'; 7477 'EPOS: Zielposition < Software-Endschalter Minus'; 7478 'EPOS: Zielposition > Software-Endschalter Plus'; 7479 'EPOS: Software-Endschalter Minus angefahren'; 7480 'EPOS: Software-Endschalter Plus angefahren'; 7481 'EPOS: Achsposition < Software-Endschalter Minus'; 7482 'EPOS: Achsposition > Software-Endschalter Plus'; 7483 'EPOS: Fahren auf Festanschlag Klemmmoment nicht erreicht'; 7484 'EPOS: Festanschlag außerhalb Überwachungsfenster'; 7485 'EPOS: Festanschlag nicht erreicht'; 7486 'EPOS: Zwischenhalt fehlt'; 7487 'EPOS: Verfahrauftrag verwerfen fehlt'; 7488 'EPOS: Relative Positionierung nicht möglich'; 7489 'EPOS: Referenzpunktkorrektur außerhalb Fenster'; 7490 'EPOS: Freigabe während Verfahren weggenommen'; 7491 'EPOS: STOP-Nocken Minus angefahren'; 7492 'EPOS: STOP-Nocken Plus angefahren'; 7493 'LR: Überlauf des Wertebereiches für Lageistwert'; 7494 'LR: Antriebsdatensatz-Umschaltung während Betrieb'; 7495 'LR: Referenzfunktion abgebrochen'; 7496 'EPOS: Freigabe nicht möglich'; 7497 'LR: Lagesetzwert aktiviert'; 7498 'LR: Messtasterauswertung nicht möglich'; 7499 'EPOS: Umkehrnocken mit falscher Verfahrrichtung angefahren'; 7503 'EPOS: STOP-Nocken mit falscher Verfahrrichtung angefahren'; 7505 'EPOS: Auftrag Festanschlag bei U/f/SLVC-Betrieb nicht möglich'; 7530 'Antrieb: Antriebsdatensatz DDS nicht vorhanden'; 7531 'Antrieb: Befehlsdatensatz CDS nicht vorhanden'; 7550 'Antrieb: Geberparameter zurücksetzen nicht möglich'; 7552 'Antrieb Geber: Geberkonfiguration nicht unterstützt'; 7553 'Antrieb Geber: Sensor Module Konfiguration nicht unterstützt'; 7557 'Geber 1: Referenzpunkt-Koordinate nicht im zulässigen Bereich'; 7558 'Geber 2: Referenzpunkt-Koordinate nicht im zulässigen Bereich'; 7563 'Antrieb Geber: XIST1_ERW Konfiguration fehlerhaft'; 7565 'Antrieb: Geberfehler PROFIdrive-Geberschnittstelle 1'; 7566 'Antrieb: Geberfehler PROFIdrive-Geberschnittstelle 2'; 7577 'Geber 1: Messtasterauswertung nicht möglich'; 7578 'Geber 2: Messtasterauswertung nicht möglich'; 7581 'Geber 1: Lageistwertaufbereitung fehlerhaft'; 7582 'Geber 2: Lageistwertaufbereitung fehlerhaft'; 7584 'Geber 1: Lagesetzwert aktiviert'; 7585 'Geber 2: Lagesetzwert aktiviert'; 7587 'Geber 1: Lageistwertaufbereitung hat keinen gültigen Geber'; 7588 'Geber 2: Lageistwertaufbereitung hat keinen gültigen Geber'; 7590 'Geber 1: Antriebsdatensatz-Umschaltung während Betrieb'; 7591 'Geber 2: Antriebsdatensatz-Umschaltung während Betrieb'; 7593 'Geber 1: Wertebereich für Lageistwert überschritten'; 7594 'Geber 2: Wertebereich für Lageistwert überschritten'; 7596 'Geber 1: Referenzfunktion abgebrochen'; 7597 'Geber 2: Referenzfunktion abgebrochen'; 7599 'Geber 1: Justage nicht möglich'; 7600 'Geber 2: Justage nicht möglich'; 7800 'Antrieb: Kein Leistungsteil vorhanden'; 7801 'Antrieb: Motor Überstrom'; 7802 'Antrieb: Einspeisung oder Leistungsteil nicht bereit'; 7805 'Antrieb: Leistungsteil Überlastung I2t'; 7806 'Antrieb: Generatorische Leistungsgrenze überschritten (F3E)'; 7807 'Antrieb: Kurzschluss/Erdschluss erkannt'; 7808 'HF Damping Module: Dämpfung nicht bereit'; 7810 'Antrieb: Leistungsteil-EEPROM ohne Nenndaten'; 7850 'Externe Warnung 1'; 7851 'Externe Warnung 2'; 7852 'Externe Warnung 3'; 7860 'Externe Störung 1'; 7861 'Externe Störung 2'; 7862 'Externe Störung 3'; 7900 'Antrieb: Motor blockiert'; 7901 'Antrieb: Motor Überdrehzahl'; 7902 'Antrieb: Motor gekippt'; 7903 'Antrieb: Motor Drehzahlabweichung'; 7910 'Antrieb: Motor Übertemperatur'; 7920 'Antrieb: Drehmoment/Drehzahl zu niedrig'; 7921 'Antrieb: Drehmoment/Drehzahl zu hoch'; 7922 'Antrieb: Drehmoment/Drehzahl außerhalb Toleranz'; 7923 'Antrieb: Drehmoment/Drehzahl zu niedrig'; 7924 'Antrieb: Drehmoment/Drehzahl zu hoch'; 7925 'Antrieb: Drehmoment/Drehzahl außerhalb Toleranz'; 7927 'Gleichstrombremsung aktiv'; 7929 'Antrieb: Kein Motor erkannt'; 7936 'Antrieb: Lastausfall'; 7950 'Motorparameter fehlerhaft'; 7967 'Antrieb: Pollageidentifikation interner Fehler'; 7968 'Antrieb: Lq-Ld-Messung fehlerhaft'; 7969 'Antrieb: Pollageidentifikation fehlerhaft'; 7975 'Antrieb: Fahren bis Nullmarke - Sollwertvorgabe erwartet'; 7976 'Antrieb: Geberfeinabgleich aktiviert'; 7980 'Antrieb: Drehende Messung aktiviert'; 7981 'Antrieb: Drehende Messung Freigaben fehlen'; 7983 'Antrieb: Drehende Messung Sättigungskennlinie'; 7984 'Antrieb: Drehzahlregleroptimierung Trägheitsmoment'; 7985 'Antrieb: Drehzahlregleroptimierung (Schwingungstest)'; 7986 'Antrieb: Drehende Messung Hochlaufgeber'; 7988 'Antrieb: Drehende Messung Keine Konfiguration ausgewählt'; 7990 'Antrieb: Motordatenidentifikation fehlerhaft'; 7991 'Antrieb: Motordatenidentifikation aktiviert'; 7994 'Antrieb: Motordatenidentifikation nicht durchgeführt'; 8010 'CU: Analog-Digital-Wandler'; 8501 'PROFINET: Sollwert Timeout'; 8502 'PROFINET: Überwachungszeit Lebenszeichen abgelaufen'; 8511 'PROFINET: Empfangs-Konfigurationsdaten ungültig'; 8526 'PROFINET: Keine zyklische Verbindung'; 8565 'PROFINET: Konsistenzfehler bei Einstellparametern'; 8760 'CAN: Überschreitung maximaler Größe des PZD IF'; 8800 'PROFIenergy Energiesparmodus aktiv'; 8802 'PROFIenergy Inkrementalgeberversorgung ausschalten nicht möglich'; 13009 'Lizenzierung OA-Applikation nicht lizenziert'; 13100 'Know-how-Schutz: Kopierschutzfehler'; 13101 'Know-how-Schutz: Kopierschutz nicht aktivierbar'; 13102 'Know-how-Schutz: Konsistenzfehler der geschützten Daten'; 30001 'Leistungsteil: Überstrom'; 30002 'Leistungsteil: Zwischenkreisspannung Überspannung'; 30003 'Leistungsteil: Zwischenkreisspannung Unterspannung'; 30004 'Leistungsteil: Übertemperatur Kühlkörper Wechselrichter'; 30005 'Leistungsteil: Überlastung I2t'; 30011 'Leistungsteil: Netzphasenausfall im Hauptstromkreis'; 30015 'Leistungsteil: Phasenausfall Motorleitung'; 30016 'Leistungsteil: Lastversorgung ausgeschaltet'; 30017 'Leistungsteil: Hardware Strombegrenzung zu oft angesprochen'; 30021 'Leistungsteil: Erdschluss'; 30022 'Leistungsteil: Überwachung U_ce'; 30024 'Leistungsteil: Übertemperatur Thermisches Modell'; 30025 'Leistungsteil: Übertemperatur Chip'; 30027 'Leistungsteil: Vorladung Zwischenkreis Zeitüberwachung'; 30031 'Leistungsteil: Hardware Strombegrenzung in Phase U'; 30032 'Leistungsteil: Hardware Strombegrenzung in Phase V'; 30033 'Leistungsteil: Hardware Strombegrenzung in Phase W'; 30034 'Leistungsteil: Übertemperatur Innenraum'; 30042 'Leistungsteil: Lüfter hat maximale Betriebsstunden erreicht'; 30052 'EEPROM Daten fehlerhaft'; 30054 'Leistungsteil: Unterspannung bei Bremse öffnen'; 30057 'Leistungsteil: Netzunsymmetrie'; 30071 'Keine neuen Istwerte von Power Module empfangen'; 30072 'Keine Sollwerte mehr an Power Module übertragbar'; 30074 'Kommunikationsfehler zwischen Control Unit und Power Module'; 30080 'Leistungsteil: Stromanstieg zu schnell'; 30081 'Leistungsteil: Schalthandlungen zu häufig'; 30105 'LT: Istwerterfassung fehlerhaft'; 30502 'Leistungsteil: Zwischenkreis Überspannung'; 30600 'SI P2: STOP A ausgelöst'; 30611 'SI P2: Defekt in einem Überwachungskanal'; 30620 'SI P2: Sicher abgeschaltetes Moment aktiv'; 30625 'SI P2: Lebenszeichen in Safety-Daten fehlerhaft'; 30649 'SI P2: Softwarefehler intern'; 30650 'SI P2: Abnahmetest erforderlich'; 30651 'SI P2: Synchronisation mit Control Unit fehlgeschlagen'; 30655 'SI P2: Abgleich der Überwachungsfunktionen'; 30656 'SI P2: Parameter Prozessor 2 fehlerhaft'; 30659 'SI P2: Schreibauftrag für Parameter abgewiesen'; 30662 'Fehler in interner Kommunikation'; 30664 'Fehler in der Hochlaufphase'; 30665 'SI P2: System ist defekt'; 30666 'SI Motion P2: Statisches 1-Signal am F-DI für sichere Quittierung'; 30680 'SI Motion P2: Prüfsummenfehler sichere Überwachungen'; 30681 'SI Motion P2: Parameterwert falsch'; 30682 'SI Motion P2: Überwachungsfunktion nicht unterstützt'; 30683 'SI Motion P2: SLS-Freigabe fehlt'; 30692 'SI Motion P2: Parameterwert falsch geberlos'; 30693 'SI P2: Safety-Parametrierung geändert POWER ON erforderlich'; 30700 'SI Motion P2: STOP A ausgelöst'; 30701 'SI Motion P2: STOP B ausgelöst'; 30706 'SI Motion P2: SAM/SBR Grenze überschritten'; 30711 'SI Motion P2: Defekt in einem Überwachungskanal'; 30712 'SI Motion P2: Defekt bei F-IO-Verarbeitung'; 30714 'SI Motion P2: Sicher begrenzte Geschwindigkeit überschritten'; 30716 'SI Motion P2: Toleranz für sichere Bewegungsrichtung überschritten'; 30770 'SI Motion P2: Diskrepanzfehler der fehlersicheren Eingänge'; 30772 'SI Motion P2: Teststop fehlersichere Eingänge/Ausgänge aktiv'; 30773 'SI Motion P2: Teststop fehlerhaft'; 30798 'SI Motion P2: Teststop läuft'; 30799 'SI Motion P2: Abnahmetestmodus aktiv'; 30800 'Leistungsteil: Sammelmeldung'; 30802 'Leistungsteil: Zeitscheibenüberlauf'; 30804 'Leistungsteil: CRC'; 30805 'Leistungsteil: Prüfsumme EPROM nicht korrekt'; 30809 'Leistungsteil: Schaltinformation ungültig'; 30810 'Leistungsteil: Watchdog Timer'; 30850 'Leistungsteil: Softwarefehler intern'; 30875 'Leistungsteil DRIVE-CLiQ (CU): Versorgungsspannung ausgefallen'; 30903 'Leistungsteil: I2C-Bus Fehler aufgetreten'; 30920 'Fehler Temperatursensor'; 30950 'Leistungsteil: Softwarefehler intern'; 30999 'Leistungsteil: Unbekannte Warnung'; 31100 'Geber 1: Nullmarkenabstand fehlerhaft'; 31101 'Geber 1: Nullmarke ausgefallen'; 31103 'Geber 1: Amplitudenfehler Spur R'; 31118 'Geber 1: Drehzahldifferenz außerhalb Toleranz'; 31131 'Geber 1: Abweichung Lage inkrementell/absolut zu groß'; 31150 'Geber 1: Initialisierung fehlerhaft'; 31400 'Geber 1: Warnschwelle Nullmarkenabstand fehlerhaft'; 31401 'Geber 1: Warnschwelle Nullmarke ausgefallen'; 31418 'Geber 1: Drehzahldifferenz je Abtastrate überschritten'; 31422 'Geber 1: Impulszahl Rechteckgeber außerhalb Toleranzband'; 31431 'Geber 1: Abweichung Lage inkrementell/absolut zu groß'; 31802 'Geber 1: Zeitscheibenüberlauf'; 31805 'Geber 1: Prüfsumme EPROM nicht 